// Mitsubishi GX Works2 project: 11国轩烘烤线体修改1028   PLC: Q06UDEH (continued)

lifter11203(ShuttleCarInOut:=LifterIO11203);(*出口升降台*)
LifterIO11203.xCylinder:=1;
Y246:=LifterIO11203.xCW;
Y247:=LifterIO11203.xCCW;
LifterIO11203.xForward:=M550;
LifterIO11203.xBackward:=M551;
ShuttleCarCurrentPosition(X51 OR X50,X50,X51,FALSE,LifterIO11203.iCurrentPos);
F455:=LifterIO11203.xOvertimeAlarm ;
LifterIO11203.diDeviceID:=11203;

Cylinder112011(ShuttleCarInOut:=	CylinderIO112011);	(*升降门*)
CylinderIO112011.xCylinder:=1;
Y240:=CylinderIO112011.xCW;(*修改*)				
Y241:=CylinderIO112011.xCCW;(*修改*)					
CylinderIO112011.xForward:=M556;				
CylinderIO112011.xBackward:=M557;				
ShuttleCarCurrentPosition(X4B OR X4A,X4B,X4A,FALSE,CylinderIO112011.iCurrentPos);				
F460:=CylinderIO112011.xOvertimeAlarm ;				
CylinderIO112011.diDeviceID:=112011;

Cylinder112012(ShuttleCarInOut:=	CylinderIO112012);	(*升降门*)
CylinderIO112012.xCylinder:=1;
Y242:=CylinderIO112012.xCW;	(*修改*)				
Y243:=CylinderIO112012.xCCW;		(*修改*)			
CylinderIO112012.xForward:=M558;				
CylinderIO112012.xBackward:=M559;				
ShuttleCarCurrentPosition(X4D OR X4C,X4D,X4C,FALSE,CylinderIO112012.iCurrentPos);				
F461:=CylinderIO112012.xOvertimeAlarm ;				
CylinderIO112012.diDeviceID:=112012;

Cylinder112041(ShuttleCarInOut:=	CylinderIO112041);	(*升降门*)
CylinderIO112041.xCylinder:=1;
Y24A:=CylinderIO112041.xCW;				
Y24B:=CylinderIO112041.xCCW;				
CylinderIO112041.xForward:=M560;				
CylinderIO112041.xBackward:=M561;				
ShuttleCarCurrentPosition(X54 OR X55,X55,X54,FALSE,CylinderIO112041.iCurrentPos);				
F462:=CylinderIO112041.xOvertimeAlarm ;				
CylinderIO112041.diDeviceID:=112041;

Cylinder112042(ShuttleCarInOut:=	CylinderIO112042);	(*升降门*)
CylinderIO112042.xCylinder:=1;
Y248:=CylinderIO112042.xCW;				
Y249:=CylinderIO112042.xCCW;				
CylinderIO112042.xForward:=M562;				
CylinderIO112042.xBackward:=M563;				
ShuttleCarCurrentPosition(X53 OR X52,X53,X52,FALSE,CylinderIO112042.iCurrentPos);				
F463:=CylinderIO112042.xOvertimeAlarm ;				
CylinderIO112042.diDeviceID:=112042;
	
Switch11301(ConveyorEntryIO:=	ConveyorIO111041,ConveyorExitIO:=	ConveyorIO11103,SwitchIO:=	SwitchIO11301);(*这里的Exit是为出线体，Entry为进线体*)
SwitchIO11301.xLiftCylinderRetractDetect:=X61;				
SwitchIO11301.xLiftCylinderExtendDetect:=X60;				
Y24C:=SwitchIO11301.xLiftCylinderExtend;				
SwitchIO11301.xLiftCylinderExtendButton:=M564;
SwitchIO11301.xLiftCylinderRetractButton:= NOT M564;		
F464:=SwitchIO11301.xOvertimeAlarm ;				

Switch11302(ConveyorEntryIO:= 	ConveyorIO111042,ConveyorExitIO:= 	ConveyorIO11106,SwitchIO:=	SwitchIO11302);
SwitchIO11302.xLiftCylinderRetractDetect:=X63;				
SwitchIO11302.xLiftCylinderExtendDetect:=X62;				
Y24D:=SwitchIO11302.xLiftCylinderExtend;				
SwitchIO11302.xLiftCylinderExtendButton:=M567;
SwitchIO11302.xLiftCylinderRetractButton:=NOT M567;				
F465:=SwitchIO11302.xOvertimeAlarm ;				

IF  m_i11315Task=1
  THEN 
 			Switch11315(ConveyorEntryIO:=ConveyorIO11137,ConveyorExitIO:=               ConveyorIO111381,	SwitchIO:= 	SwitchIO11315 );
   ELSE
     		Switch11315(ConveyorEntryIO:=ConveyorIO111381,ConveyorExitIO:=               ConveyorIO11137,	SwitchIO:= 	SwitchIO11315 );
END_IF;
SwitchIO11315.xLiftCylinderRetractDetect:=X7D;				
SwitchIO11315.xLiftCylinderExtendDetect:=X7C;				
Y25A:=SwitchIO11315.xLiftCylinderExtend;				
Y266:=SwitchIO11315.xEntryBarCylinderRetract;				
Y260:=(g_xAuto AND  m_i11315Task=2 )OR (M720 AND g_xManual) ;	(*十字路口阻挡气缸输出1*)	
Y261:=(g_xAuto AND  m_i11315Task=1 )OR ( M721 AND g_xManual);	(*十字路口阻挡气缸输出2*)
SwitchIO11315.xLiftCylinderExtendButton:=M568;	
SwitchIO11315.xLiftCylinderRetractButton:= NOT M568;	
SwitchIO11315.xEntryBarCylinderRetractButton:=M569;				
SwitchIO11315.xExitBarCylinderRetractButton:=M570;				
F466:=SwitchIO11315.xOvertimeAlarm ;				

Switch11316(ConveyorEntryIO:=ConveyorIO11140,ConveyorExitIO:= 	ConveyorIO111382,SwitchIO:= 	SwitchIO11316 );
SwitchIO11316.xLiftCylinderRetractDetect:=X7F;				
SwitchIO11316.xLiftCylinderExtendDetect:=X7E;				
Y25B:=SwitchIO11316.xLiftCylinderExtend;				
Y268:=NOT (m_i11316Task=2 OR M722);(*316阻挡气缸1*)		
Y269:=NOT (m_i11316Task=1 OR M723);	(*316阻挡气缸2*)	
SwitchIO11316.xLiftCylinderExtendButton:=M571;
SwitchIO11316.xLiftCylinderRetractButton:= NOT M571;				
SwitchIO11316.xEntryBarCylinderRetractButton:=M572;				
F467:=SwitchIO11316.xOvertimeAlarm ;				

UConveyor11303(	ConveyorIOLeft:=ConveyorIO11118,	ConveyorIORight:=ConveyorIO11120,	
									ConveyorIODown:=ConveyorIO11113,	UConveyorIO:=UConveyorIO11303);
UConveyorIO11303.xLiftCylinderExtendDetect1:=X64;
UConveyorIO11303.xLiftCylinderRetractDetect1:=X65;									
Y24E:=UConveyorIO11303.xLiftCylinderExtend1;								
Y262:=UConveyorIO11303.xExitBarCylinderRetract1;								
UConveyorIO11303.xLiftCylinderRetractDetect2:=X69;								
UConveyorIO11303.xLiftCylinderExtendDetect2:=X68;		
UConveyorIO11303.xBatteryDetect1:=X1A;		
Y250:=UConveyorIO11303.xLiftCylinderExtend2;								
UConveyorIO11303.xLiftCylinderExtendButton1:=M573;								
UConveyorIO11303.xExitBarCylinderRetractButton1:=M574;								
UConveyorIO11303.xLiftCylinderExtendButton2:=M575;								
F468:=UConveyorIO11303.xOvertimeAlarm ;								
(**X1A为电池检测保护*)

UConveyor11306(	ConveyorIOLeft:=ConveyorIO11121,	ConveyorIORight:=ConveyorIO11123,	
									ConveyorIODown:=ConveyorIO11114,	UConveyorIO:=UConveyorIO11306);
UConveyorIO11306.xLiftCylinderExtendDetect1:=X6A;	
UConveyorIO11306.xLiftCylinderRetractDetect1:=X6B;		
UConveyorIO11306.xBatteryDetect1:=X1F;							
Y251:=UConveyorIO11306.xLiftCylinderExtend1;								
Y263:=  UConveyorIO11306.xExitBarCylinderRetract1 ;								
UConveyorIO11306.xLiftCylinderRetractDetect2:=X6F;								
UConveyorIO11306.xLiftCylinderExtendDetect2:=X6E;								
Y253:=UConveyorIO11306.xLiftCylinderExtend2;								
UConveyorIO11306.xLiftCylinderExtendButton1:=M576;								
UConveyorIO11306.xExitBarCylinderRetractButton1:=M577;								
UConveyorIO11306.xLiftCylinderExtendButton2:=M578;								
F469:=UConveyorIO11306.xOvertimeAlarm ;								
(**X1F为电池检测保护*)

UConveyor11309(	ConveyorIOLeft:=ConveyorIO11124,	ConveyorIORight:=ConveyorIO11126,	
									ConveyorIODown:=ConveyorIO11115,	UConveyorIO:=UConveyorIO11309);
UConveyorIO11309.xLiftCylinderExtendDetect1:=X70;	
UConveyorIO11309.xLiftCylinderRetractDetect1:=X71;							
Y254:=UConveyorIO11309.xLiftCylinderExtend1;								
Y264:=UConveyorIO11309.xExitBarCylinderRetract1;								
UConveyorIO11309.xLiftCylinderRetractDetect2:=X75;								
UConveyorIO11309.xLiftCylinderExtendDetect2:=X74;								
Y256:=UConveyorIO11309.xLiftCylinderExtend2;								
UConveyorIO11309.xLiftCylinderExtendButton1:=M579;								
UConveyorIO11309.xExitBarCylinderRetractButton1:=M580;								
UConveyorIO11309.xLiftCylinderExtendButton2:=M581;								
F470:=UConveyorIO11309.xOvertimeAlarm ;								
(**X22为电池检测保护*)

UConveyor11312(	ConveyorIOLeft:=ConveyorIO11127,	ConveyorIORight:=ConveyorIO11129,	
									ConveyorIODown:=ConveyorIO11116,	UConveyorIO:=UConveyorIO11312);
UConveyorIO11312.xLiftCylinderExtendDetect1:=X76;
UConveyorIO11312.xLiftCylinderRetractDetect1:=X77;								
Y257:=UConveyorIO11312.xLiftCylinderExtend1;								
Y265:=UConveyorIO11312.xExitBarCylinderRetract1;								
UConveyorIO11312.xLiftCylinderRetractDetect2:=X7B;								
UConveyorIO11312.xLiftCylinderExtendDetect2:=X7A;								
Y259:=UConveyorIO11312.xLiftCylinderExtend2;								
UConveyorIO11312.xLiftCylinderExtendButton1:=M582;								
UConveyorIO11312.xExitBarCylinderRetractButton1:=M583;								
UConveyorIO11312.xLiftCylinderExtendButton2:=M584;								
F471:=UConveyorIO11312.xOvertimeAlarm ;								

(**************通信地址分配***************)
ComConveyor11104(ConveyorIO:=ConveyorIO11104,CommunicationIO:=ComConveyorIO11104);
ComCOnveyorIO11104.i_iResponsPCPLC:=D2001;	
ComCOnveyorIO11104.i_iReadWriteFlagPCPLC:=D2006;	
ComCOnveyorIO11104.i_iTaskProcessFlagPCPLC:=D2007;	
ComCOnveyorIO11104.i_iCommandPCPLC:=D2008;	
ComCOnveyorIO11104.i_iTaskIDPCPLC:=D2009;	
DMOV(TRUE,D2010,ComConveyorIO11104.i_diDestinationDevicePCPLC);	
ComCOnveyorIO11104.i_iProductIDPCPLC:=D2012;	
D3001:=ComCOnveyorIO11104.o_iRequestPLCPC;	
D3006:=ComCOnveyorIO11104.o_iReadWriteFlagPLCPC;	
D3007:=ComCOnveyorIO11104.o_iDeviceStatusPLCPC;	
D3008:=ComCOnveyorIO11104.o_iTaskIDPLCPC;	
D3009:=ComCOnveyorIO11104.o_iProductIDPLCPC;	

ComConveyor11108(ConveyorIO:=ConveyorIO11108,CommunicationIO:=ComConveyorIO11108);
ComCOnveyorIO11108.i_iResponsPCPLC:=D2016;	
ComCOnveyorIO11108.i_iReadWriteFlagPCPLC:=D2021;	
ComCOnveyorIO11108.i_iTaskProcessFlagPCPLC:=D2022;	
ComCOnveyorIO11108.i_iCommandPCPLC:=D2023;	
ComCOnveyorIO11108.i_iTaskIDPCPLC:=D2024;	
DMOV(TRUE,D2025,ComConveyorIO11108.i_diDestinationDevicePCPLC);		
ComCOnveyorIO11108.i_iProductIDPCPLC:=D2027;	
D3016:=ComCOnveyorIO11108.o_iRequestPLCPC;	
D3021:=ComCOnveyorIO11108.o_iReadWriteFlagPLCPC;	
D3022:=ComCOnveyorIO11108.o_iDeviceStatusPLCPC;	
D3023:=ComCOnveyorIO11108.o_iTaskIDPLCPC;	
D3024:=ComCOnveyorIO11108.o_iProductIDPLCPC;	

ComConveyor11107(ConveyorIO:=ConveyorIO11107,CommunicationIO:=ComConveyorIO11107);
ComConveyorIO11107.i_iResponsPCPLC:=D2031;	
ComConveyorIO11107.i_iReadWriteFlagPCPLC:=D2036;	
ComConveyorIO11107.i_iTaskProcessFlagPCPLC:=D2037;	
ComConveyorIO11107.i_iCommandPCPLC:=D2038;	
ComConveyorIO11107.i_iTaskIDPCPLC:=D2039;	
DMOV(TRUE,D2040,ComConveyorIO11107.i_diDestinationDevicePCPLC);	
ComConveyorIO11107.i_iProductIDPCPLC:=D2042;	
D3031:=ComConveyorIO11107.o_iRequestPLCPC;	
D3036:=ComConveyorIO11107.o_iReadWriteFlagPLCPC;	
D3037:=ComConveyorIO11107.o_iDeviceStatusPLCPC;	
D3038:=ComConveyorIO11107.o_iTaskIDPLCPC;	
D3039:=ComConveyorIO11107.o_iProductIDPLCPC;	
	

ComConveyor11142(ConveyorIO:=ConveyorIO11142,CommunicationIO:=ComConveyorIO11142);
ComCOnveyorIO11142.i_iResponsPCPLC:=D2046;	
ComCOnveyorIO11142.i_iReadWriteFlagPCPLC:=D2051;	
ComCOnveyorIO11142.i_iTaskProcessFlagPCPLC:=D2052;	
ComCOnveyorIO11142.i_iCommandPCPLC:=D2053;	
ComCOnveyorIO11142.i_iTaskIDPCPLC:=D2054;	
DMOV(TRUE,D2055,ComConveyorIO11142.i_diDestinationDevicePCPLC);	
ComCOnveyorIO11142.i_iProductIDPCPLC:=D2057;	
D3046:=ComCOnveyorIO11142.o_iRequestPLCPC;	
D3051:=ComCOnveyorIO11142.o_iReadWriteFlagPLCPC;	
D3052:=ComCOnveyorIO11142.o_iDeviceStatusPLCPC;	
D3053:=ComCOnveyorIO11142.o_iTaskIDPLCPC;	
D3054:=ComCOnveyorIO11142.o_iProductIDPLCPC;	

ComConveyor11141(ConveyorIO:=ConveyorIO11141,CommunicationIO:=ComConveyorIO11141);
ComCOnveyorIO11141.i_iResponsPCPLC:=D2061;	
ComCOnveyorIO11141.i_iReadWriteFlagPCPLC:=D2066;	
ComCOnveyorIO11141.i_iTaskProcessFlagPCPLC:=D2067;	
ComCOnveyorIO11141.i_iCommandPCPLC:=D2068;	
ComCOnveyorIO11141.i_iTaskIDPCPLC:=D2069;	
DMOV(TRUE,D2070,ComConveyorIO11141.i_diDestinationDevicePCPLC);	
ComCOnveyorIO11141.i_iProductIDPCPLC:=D2072;	
D3061:=ComCOnveyorIO11141.o_iRequestPLCPC;	
D3066:=ComCOnveyorIO11141.o_iReadWriteFlagPLCPC;	
D3067:=ComCOnveyorIO11141.o_iDeviceStatusPLCPC;	
D3068:=ComCOnveyorIO11141.o_iTaskIDPLCPC;	
D3069:=ComCOnveyorIO11141.o_iProductIDPLCPC;	

ComConveyor11110(ConveyorIO:=ConveyorIO11110,CommunicationIO:=ComConveyorIO11110);
ComCOnveyorIO11110.i_iResponsPCPLC:=D2076;	
ComCOnveyorIO11110.i_iReadWriteFlagPCPLC:=D2081;	
ComCOnveyorIO11110.i_iTaskProcessFlagPCPLC:=D2082;	
ComCOnveyorIO11110.i_iCommandPCPLC:=D2083;	
ComCOnveyorIO11110.i_iTaskIDPCPLC:=D2084;	
DMOV(TRUE,D2085,ComConveyorIO11110.i_diDestinationDevicePCPLC);	
ComCOnveyorIO11110.i_iProductIDPCPLC:=D2087;	
D3076:=ComCOnveyorIO11110.o_iRequestPLCPC;	
D3081:=ComCOnveyorIO11110.o_iReadWriteFlagPLCPC;	
D3082:=ComCOnveyorIO11110.o_iDeviceStatusPLCPC;	
D3083:=ComCOnveyorIO11110.o_iTaskIDPLCPC;	
D3084:=ComCOnveyorIO11110.o_iProductIDPLCPC;	

ComConveyor11111(ConveyorIO:=ConveyorIO11111,CommunicationIO:=ComConveyorIO11111);
ComCOnveyorIO11111.i_iResponsPCPLC:=D2091;	
ComCOnveyorIO11111.i_iReadWriteFlagPCPLC:=D2096;	
ComCOnveyorIO11111.i_iTaskProcessFlagPCPLC:=D2097;	
ComCOnveyorIO11111.i_iCommandPCPLC:=D2098;	
ComCOnveyorIO11111.i_iTaskIDPCPLC:=D2099;	
DMOV(TRUE,D2100,ComConveyorIO11111.i_diDestinationDevicePCPLC);	
ComCOnveyorIO11111.i_iProductIDPCPLC:=D2102;	
D3091:=ComCOnveyorIO11111.o_iRequestPLCPC;	
D3096:=ComCOnveyorIO11111.o_iReadWriteFlagPLCPC;	
D3097:=ComCOnveyorIO11111.o_iDeviceStatusPLCPC;	
D3098:=ComCOnveyorIO11111.o_iTaskIDPLCPC;	
D3099:=ComCOnveyorIO11111.o_iProductIDPLCPC;	

ComConveyor11143(ConveyorIO:=ConveyorIO11143,CommunicationIO:=ComConveyorIO11143);
ComConveyorIO11143.i_iResponsPCPLC:=D2106;	
ComConveyorIO11143.i_iReadWriteFlagPCPLC:=D2111;	
ComConveyorIO11143.i_iTaskProcessFlagPCPLC:=D2112;	
ComConveyorIO11143.i_iCommandPCPLC:=D2113;	
ComConveyorIO11143.i_iTaskIDPCPLC:=D2114;	
DMOV(TRUE,D2115,ComConveyorIO11143.i_diDestinationDevicePCPLC);	
ComConveyorIO11143.i_iProductIDPCPLC:=D2117;	
D3106:=ComConveyorIO11143.o_iRequestPLCPC;	
D3111:=ComConveyorIO11143.o_iReadWriteFlagPLCPC;	
D3112:=ComConveyorIO11143.o_iDeviceStatusPLCPC;	
D3113:=ComConveyorIO11143.o_iTaskIDPLCPC;	
D3114:=ComConveyorIO11143.o_iProductIDPLCPC;	

(*///////////////////////////////////自动部分/////////////////////////////*)
IF g_xAuto    THEN
			(*门直接用Y控制，不用块了*)
			CylinderIO112011.xMDIExe:=1;
		IF D401.2  AND 	ConveyorIO11101.xEmpty  AND CylinderIO112012.iCurrentPos=1
			THEN(*上层10给11有料信号401.2*)
						CylinderIO112011.iDestinationPos:=2;
			ELSE CylinderIO112011.iDestinationPos:=1; (*如果10有下料信号但是11对接线体也有料，则关闭AB门*)
		END_IF;	
		D201.2:=CylinderIO112011.iCurrentPos=2 AND ConveyorIO11101.xEmpty;(*11给10的上层下料允许对接信号*)
		ConveyorIO11101.xLoad:=D401.4;(*10线体的下料信号*)
		(*第2个隔离门*)
		CylinderIO112012.xMDIExe:=1;
		IF NOT ConveyorIO11101.xEmpty  AND CylinderIO112011.iCurrentPos=1 (*第二个隔离门只有在第一个隔离门关住后*)
			THEN
							CylinderIO112012.iDestinationPos:=2;
			ELSE 	CylinderIO112012.iDestinationPos:=1;
		END_IF;		
		ConveyorIO11101.xUnload:=ConveyorIO11102.xEmpty AND CylinderIO112012.iCurrentPos=2;
		ConveyorIO11102.xLoad:=ConveyorIO11101.xNextRun;
		Switch11301Task(xCondition:= Switch11301Condition,(*抢占排队*)
									xTaskComplete:=LDP(TRUE,ConveyorIO111041.xEmpty) ,
									xReset:=g_diDeviceIDSelect=11104 AND g_xResetSingle ,
									iPriority:=m_i11301Task);
		Switch11301Condition[1]:=ConveyorIO11102.xEmpty=0 AND ConveyorIO11104.xEmpty;(*顶升移栽任务1,往烘烤*)
		Switch11301Condition[2]:=ConveyorIO11109.xEmpty=0 AND ConveyorIO11111.xEmpty AND LifterIO11202.iCurrentPos=2;(*顶升移栽任务2，往机械手*)
		ConveyorIO11102.xUnload:=ConveyorIO111041.xEmpty AND m_i11301Task=1;
		SwitchIO11301.xLiftCylinderExtendInit:=1;(*初始化顶起*)
		SwitchIO11301.xEntryEnable:=ConveyorIO11102.xNextRun;
		SwitchIO11301.xSwithEnable:=m_i11301Task=2;(*任务2要直行，降下气缸*)
		SwitchIO11301.xExitEnable:=(ConveyorIO11104.xEmpty AND m_i11301Task=1)(*1041虚拟线体运给104*)
													OR(ConveyorIO11111.xEmpty AND m_i11301Task=2);(*11103出料给11111*)
		(*满框去烘烤*)													
		ConveyorIO11104.xLoad:=ConveyorIO111041.xNextRun;
		ConveyorIO11104.xUnload:=ConveyorIO111042.xEmpty;(*这里到时候需要加一个扫码条件，判断去哪个烘烤库*)
		SwitchIO11302.xEntryEnable:=ConveyorIO11104.xNextRun;
		SwitchIO11302.xSwithEnable:=1;
		SwitchIO11302.xLiftCylinderExtendInit:=1;(*初始化顶起*)
		SwitchIO11302.xExitEnable:=(ConveyorIO111042.diDesConveyor=11108 AND ConveyorIO11108.xEmpty)
													OR (ConveyorIO111042.diDesConveyor=11107 AND ConveyorIO11107.xEmpty);
		ConveyorIO11106.xUnloadCCW:=ConveyorIO111042.diDesConveyor=11108;
		ConveyorIO11107.xLoad:=ConveyorIO11106.xNextRun AND  ConveyorIO11106.diDesConveyor=11107;
		ConveyorIO11108.xLoad:=ConveyorIO11106.xNextRun AND ConveyorIO11106.diDesConveyor=11108;
		(*未增加11107和11108下料信号，与工控机信号对接*)
		Switch11316Task(arrxCondition:=Switch11316Condition ,
								xTaskComplete:= LDF(TRUE,ConveyorIO11138.xEmpty),
								xReset:= g_xResetSingle AND g_diDeviceIDSelect=11138,	
								iPriority:=m_i11316Task);
		Switch11316Condition[1].xCondition:=ConveyorIO11141.xEmpty=0;
		Switch11316Condition[2].xCondition:=ConveyorIO11142.xEmpty=0;
		
		LifterIO11204.xMDIExe:=NOT ConveyorIO11140.xError AND NOT ConveyorIO11141.xError ;
		IF NOT ConveyorIO11142.xEmpty   THEN
			LifterIO11204.iDestinationPos:=1;
		ELSE 
			LifterIO11204.iDestinationPos:=2;
		END_IF;	

		LifterIO11205.xMDIExe:=NOT ConveyorIO11140.xError AND NOT ConveyorIO11142.xError ;
		IF NOT ConveyorIO11141.xEmpty THEN
			LifterIO11205.iDestinationPos:=1;
		ELSE
			LifterIO11205.iDestinationPos:=2;
		END_IF;	
		
		(*ConveyorIO11141.xPutInto:=  M880;*)(*这里需要上位机给命令，以后需要就加*)
	(*	ConveyorIO11142.xPutInto:=  M881;*)(*这里需要上位机给命令，以后需要就加*)
		ConveyorIO11141.xUnload:=ConveyorIO11140.xEmpty AND m_i11316Task=1 ; (*AND LifterIO11204.iCurrentPos=1;*)(*这里可能需要Load，接到堆垛机指令就Load，以后需要就加*)
		ConveyorIO11142.xUnload:=ConveyorIO11140.xEmpty AND m_i11316Task=2;(*  AND LifterIO11205.iCurrentPos=1;*)
		SwitchIO11316.xEntryEnable:=(ConveyorIO11141.xNextRun AND m_i11316Task=1)
													OR (ConveyorIO11142.xNextRun AND m_i11316Task=2);
		ConveyorIO11140.xloadCCW:= m_i11316Task=1;													
		SwitchIO11316.xSwithEnable:=1;
		SwitchIO11316.xExitEnable:=ConveyorIO11138.xEmpty;
		(*下层十字路口——+——+——+——+——+——+——+——+——+——+*)
		Switch11315Task(xCondition:=Switch11315Condition ,
									xTaskComplete:=LDF(TRUE,(ConveyorIO11109.xEmpty AND m_i11315Task=2 )OR(ConveyorIO11143.xEmpty AND m_i11315Task=1) ),
									xReset:=g_xResetSingle AND g_diDeviceIDSelect=11138 ,
									iPriority:= m_i11315Task );
		Switch11315Condition[1]:=ConveyorIO11136.xEmpty=0 AND ConveyorIO11143.xEmpty;
		Switch11315Condition[2]:=(ConveyorIO11140.xEmpty=0 OR ConveyorIO111382.xEmpty=0) AND ConveyorIO11109.xEmpty AND LifterIO11202.iCurrentPos=1;(*像这种带位置判断的，最好把检测开关也加上去*)
		SwitchIO11315.xEntryEnable:=ConveyorIO11136.xNextRun OR ConveyorIO11138.xNextRun ;
		SwitchIO11315.xSwithEnable:=(*m_i11315Task=1 *)1 ;
		SwitchIO11315.xExitEnable:=(m_i11315Task=1 AND  ConveyorIO11143.xEmpty)
													OR (m_i11315Task=2 AND ConveyorIO11109.xEmpty AND  LifterIO11202.iCurrentPos=1);
		ConveyorIO11138.xload:=ConveyorIO111382.xNextRun;
		ConveyorIO11138.xUnload:=ConveyorIO111381.xEmpty AND m_i11315Task=2 AND SwitchIO11315.xLiftCylinderExtendDetect  ;
		ConveyorIO11109.xLoad:=ConveyorIO11137.xNextRun AND m_i11315Task =2;

		IF m_i11315Task=2 THEN(*任务2时，升降由11137的状态控制，1时会由Switch块自己控制。因为任务2时，走134的step,不会控制升降*)
(*			IF NOT ConveyorIO11138.xEmpty THEN
				SwitchIO11315.xLiftCylinderExtend:=1;
				SwitchIO11315.xLiftCylinderRetract:=0;
			ELSE
				SwitchIO11315.xLiftCylinderExtend:=0;
				SwitchIO11315.xLiftCylinderRetract:=1;	
			END_IF;*)
			SwitchIO11315.xLiftCylinderExtendInit:=1;
		ELSE
			SwitchIO11315.xLiftCylinderExtendInit:=0;
		END_IF;
	

		IF LDP(TRUE,NOT ConveyorIO111381.xEmpty )THEN(*原来136和137公用一个光电检测开关，137竖向，136横向，当137有料时136也有料，这里用来给136直接下料，修改后用于1381虚拟线体和137线体*)
	ConveyorIO11137.xPutInto:=1;
		ELSIF	 LDP(TRUE,NOT ConveyorIO11137.xEmpty )THEN
			ConveyorIO11137.xPutInto:=0;
		END_IF;	

													
(*11202升降控制*)
													
		LifterIO11202.xMDIExe:=NOT ConveyorIO11109.xError AND NOT ConveyorIO11103.xError AND NOT ConveyorIO11137.xError;
		ConveyorIO11109.xloadCCW:=1;
		IF ConveyorIO11109.xEmpty THEN
			LifterIO11202.iDestinationPos:=1;
		ELSE
			LifterIO11202.iDestinationPos:=2;
		END_IF;	
		IF m_i11301Task=2 THEN
		SwitchIO11301.xLiftCylinderExtend:=0;
		SwitchIO11301.xLiftCylinderRetract:=1;
		END_IF;	 
		ConveyorIO11109.xUnload:=ConveyorIO11103.xEmpty AND LifterIO11202.iCurrentPos=2 AND m_i11301Task=2;
		ConveyorIO11103.xLoad:=ConveyorIO11109.xNextRun;
		IF LDP(TRUE,ConveyorIO11103.xEmpty=0) AND m_i11301Task=2 THEN
			ConveyorIO111041.xPutInto:=1;
		ELSIF LDP(TRUE,ConveyorIO111041.xEmpty=0) AND m_i11301Task=2 THEN
			ConveyorIO111041.xPutInto:=0;	
		END_IF;
		(*烘烤出去机械手*)
		ConveyorIO11111.xLoad:=ConveyorIO11103.xNextRun;
		ConveyorIO11111.xUnload:=ConveyorIO11112.xEmpty;
		ConveyorIO11112.xLoad:=ConveyorIO11111.xNextRun;
		ConveyorIO11112.xUnload:=ConveyorIO11105.xEmpty;
		ConveyorIO11105.xLoad:=ConveyorIO11112.xNextRun;
		ConveyorIO11105.xUnload:=ConveyorIO11139.xEmpty;
		ConveyorIO11139.xLoad:=ConveyorIO11105.xNextRun;
		ConveyorIO11139.xUnload:=UConveyorio11303.iTask=1 AND m_xU1TaskStart;(*39下料给U1*)


		Conveyor11139Task(arrxCondition:=Conveyor11139Condition,
											xTaskComplete:=LDP(TRUE,ConveyorIO11139.xEmpty),
											xReset:= g_xResetSingle AND g_diDeviceIDSelect=11139 ,
											iPriority:= m_i11139Task);
		Conveyor11139Condition[1].xCondition:=ConveyorIO111181.xEmpty AND m_xLoadPermit1;
		Conveyor11139Condition[2].xCondition:=ConveyorIO111231.xEmpty  AND m_xLoadPermit2;
		Conveyor11139Condition[3].xCondition:=ConveyorIO111241.xEmpty  AND m_xLoadPermit3;
		Conveyor11139Condition[4].xCondition:=ConveyorIO111291.xEmpty  AND m_xLoadPermit4; 
		DMOV(m_i11139Task=1,	11118,	ConveyorIO11139.diDesConveyor);(*上电时，机械手U型线体处空时生成任务号，并进行抢占*)
		DMOV(m_i11139Task=2,	11123,	ConveyorIO11139.diDesConveyor);
		DMOV(m_i11139Task=3,	11124,	ConveyorIO11139.diDesConveyor);
		DMOV(m_i11139Task=4,	11129,	ConveyorIO11139.diDesConveyor);

		(*这个PickDone信号，他们给信号时置位，为empty的上升沿复位*)
		SET(XA0	AND NOT ConveyorIO11119.xEmpty,	m_xPickDone[1]);	
		RST(ConveyorIO11119.xEmpty,	m_xPickDone[1]);
		SET(XA1 	AND NOT ConveyorIO11122.xEmpty,	m_xPickDone[2]);	
		RST(ConveyorIO11122.xEmpty,	m_xPickDone[2]);
		SET(XA2	AND NOT ConveyorIO11125.xEmpty,	m_xPickDone[3]);	
		RST(ConveyorIO11125.xEmpty,	m_xPickDone[3]);
		SET(XA3	AND NOT ConveyorIO11128.xEmpty,	m_xPickDone[4]);	
		RST(ConveyorIO11128.xEmpty,	m_xPickDone[4]);

		DMOV(m_xPickDone[1] AND ConveyorIO11145.xEmpty AND ConveyorIO11145.diDesConveyor=0,	11117,	ConveyorIO11145.diDesConveyor);(*机械手给空框完成信号后将提升机线体作为目标地址发送，空框一直送至11117*)
		DMOV(m_xPickDone[2] AND ConveyorIO11146.xEmpty AND ConveyorIO11146.diDesConveyor=0,	11117,	ConveyorIO11146.diDesConveyor);
		DMOV(m_xPickDone[3] AND ConveyorIO11147.xEmpty AND ConveyorIO11147.diDesConveyor=0,	11117,	ConveyorIO11147.diDesConveyor);
		DMOV(m_xPickDone[4],	11117,	ConveyorIO11128.diDesConveyor);(*最初始的目标地址生成,*)

		(*目标地址的传递，横纵传递分开写，横纵之间的传递在块里写好了，不用担心*)
		ConveyorIO11113.diDesConveyorIn:=	ConveyorIO11139.diDesConveyorOut;
		ConveyorIO11145.diDesConveyorIn:=	ConveyorIO11113.diDesConveyorOut;
		ConveyorIO11114.diDesConveyorIn:=	ConveyorIO11145.diDesConveyorOut;
		ConveyorIO11146.diDesConveyorIn:=	ConveyorIO11114.diDesConveyorOut;
		ConveyorIO11115.diDesConveyorIn:=	ConveyorIO11146.diDesConveyorOut;
		ConveyorIO11147.diDesConveyorIn:=	ConveyorIO11115.diDesConveyorOut;
		ConveyorIO11116.diDesConveyorIn:=	ConveyorIO11147.diDesConveyorOut;
		(*纵向任务传递，包括虚拟线体*)
		ConveyorIO11120.diDesConveyorIn:=	ConveyorIO11119.diDesConveyorOut;
		ConveyorIO11121.diDesConveyorIn:=	ConveyorIO11122.diDesConveyorOut;
		ConveyorIO11126.diDesConveyorIn:=	ConveyorIO11125.diDesConveyorOut;
		ConveyorIO11127.diDesConveyorIn:=	ConveyorIO11128.diDesConveyorOut;
		ConveyorIO111042.diDesConveyor:=11107;


		m_TPU1TaskComplete(IN:=ConveyorIO11113.xEmpty ,PT:=t#200ms,Q:= m_xU1TaskComplete,ET:= m_tU1TaskComplete );
		m_TonU1TaskStart(IN:= ConveyorIO11113.xEmpty ,PT:= t#300MS ,Q:=m_xU1TaskStart ,ET:=m_tU1TaskStart );
		Uconveyor11303Task(xCondition:=Uconveyor11303Condition,
											xTaskComplete:=LDF(TRUE,m_xU1TaskComplete) ,
											xReset:= g_xResetSingle AND g_diDeviceIDSelect=11113 ,
											iPriority:=UConveyorio11303.iTask );
			Uconveyor11303Condition[1]:=ConveyorIO11139.xEmpty=0 AND m_i11139Task>0;(*这里还要再改的*)(*任务1是U块入料到机械手*)
			Uconveyor11303Condition[3]:=ConveyorIO111201.xEmpty=0  AND m_xPickDone[1];	(*任务3是右臂出料*)
		UConveyorio11303.xEntryEnable1:=ConveyorIO11139.xNextRun;(*U型横向线体入料使能，EntryEnable1，2，3都是在任务1时用*)
		UConveyorIO11303.xEntryEnable3:=ConveyorIO111201.xNextRun;(*U型右臂入料使能*)
		UConveyorio11303.xExitEnable1:=ConveyorIO11145.xEmpty ;(*xExitEnable1是主线体出，2是左臂出，3是右臂出，这个为横向线体出料使能*)
		UConveyorio11303.xExitEnable3:=ConveyorIO111181.xEmpty;(*这个为右臂出料使能*)
	
		ConveyorIO111181.xLoad:=ConveyorIO11118.xNextRun;(*这里是U块左右臂再增加一段线体时使用，用于控制该线体*)
		IF ConveyorIO111181.xEmpty=0  AND ConveyorIO11119.xEmpty THEN
			UConveyorIO11303.xLiftCylinderExtend2:=0;
			UConveyorIO11303.xLiftCylinderRetract2:=1;(*Extend2和Retract2为右臂顶升移栽气缸伸出和收回，Extend1和Retract1为左臂顶升移栽气缸伸出和收回*)
		END_IF;	
		ConveyorIO111181.xUnload:=ConveyorIO11119.xEmpty AND UConveyorIO11303.xLiftCylinderRetractDetect1 AND UConveyorIO11303.xLiftCylinderRetractDetect2;(*机械手横向线体控制*)
		ConveyorIO11119.xLoad:=ConveyorIO111181.xNextRun AND UConveyorIO11303.xLiftCylinderRetractDetect1 AND UConveyorIO11303.xLiftCylinderRetractDetect1;
			m_Ton11119(IN:= NOT ConveyorIO11119.xEmpty,PT:= t#3s ,Q:= m_x111201 ,ET:= m_t111201);
		IF NOT ConveyorIO11119.xEmpty AND m_x111201 THEN(*需加延时刷新111201，线体第0步要延时100ms才能检测有料，*)
			ConveyorIO111201.xPutInto:=1;
		ELSE 
			ConveyorIO111201.xPutInto:=0;
		END_IF;	
		ConveyorIO111201.xUnload:=ConveyorIO11120.xEmpty AND UConveyorio11303.iTask=3 ;(*右臂出料*)
	(**)	
		ConveyorIO11120.xLoadCCW:=1;
(*	 UConveyorIO11303.	xLiftCylinderExtendInit1=1 *)
		(*至此，U1的动作全部完成*)
		(*过度线体145*)
		ConveyorIO11145.xLoad:=ConveyorIO11113.xNextRun;
		ConveyorIO11145.xUnload:=(UConveyorio11306.iTask=1  AND m_xU2TaskStart )OR (ConveyorIO11146.diDesConveyor=11117 AND ConveyorIO11115.xEmpty) ;
		(*U2块*)
		m_TPU2TaskComplete(IN:=ConveyorIO11114.xEmpty ,PT:=t#200ms,Q:= m_xU2TaskComplete,ET:= m_tU2TaskComplete );
		m_TonU2TaskStart(IN:= ConveyorIO11114.xEmpty ,PT:= t#300MS ,Q:=m_xU2TaskStart ,ET:=m_tU2TaskStart );
		Uconveyor11306Task(xCondition:=Uconveyor11306Condition,
											xTaskComplete:=LDF(TRUE,m_xU2TaskComplete) ,
											xReset:= g_xResetSingle AND g_diDeviceIDSelect=11114,
											iPriority:=UConveyorIO11306.iTask );
			Uconveyor11306Condition[1]:=ConveyorIO11145.xEmpty=0 AND ConveyorIO11145.diDesConveyor<>11118
																														AND ConveyorIO11145.diDesConveyor<>0;(*这里还要再改的*)
			Uconveyor11306Condition[2]:=ConveyorIO111211.xEmpty=0  AND m_xPickDone[2];(*任务2是左臂出料*)
		UConveyorio11306.xEntryEnable1:=ConveyorIO11145.xNextRun ;
		UConveyorIO11306.xEntryEnable2:=ConveyorIO111211.xNextRun;
		UConveyorio11306.xExitEnable1:=ConveyorIO11146.xEmpty ;(*U型块任务1都是进前判断3个任务：往左进，往右进，主线体直接走，2是往左臂线体出，3是往右臂线体出*)
		UConveyorio11306.xExitEnable2:=ConveyorIO111231.xEmpty;(*xExitEnable1是主线体出，2是左臂出，3是右臂出*)
		ConveyorIO111231.xLoad:=ConveyorIO11123.xNextRun;

		IF ConveyorIO111231.xEmpty=0  AND ConveyorIO11122.xEmpty THEN
			UConveyorIO11306.xLiftCylinderExtend1:=0;
			UConveyorIO11306.xLiftCylinderRetract1:=1;(*U1,U3用2，U2,U4用1*)
		END_IF;	
		ConveyorIO111231.xUnload:=ConveyorIO11122.xEmpty AND UConveyorIO11306.xLiftCylinderRetractDetect1 AND UConveyorIO11306.xLiftCylinderRetractDetect2;(*机械手横向线体控制*)
		ConveyorIO11122.xLoad:=ConveyorIO111231.xNextRun AND UConveyorIO11306.xLiftCylinderRetractDetect1 AND UConveyorIO11306.xLiftCylinderRetractDetect2;
		m_Ton11122(IN:= NOT ConveyorIO11122.xEmpty,PT:= t#3s ,Q:= m_x111211 ,ET:= m_t111211);
		IF NOT ConveyorIO11122.xEmpty AND m_x111211 THEN(*加延时刷新111211，线体第0步要延时100ms才能检测有料，*)
			ConveyorIO111211.xPutInto:=1;
		ELSIF ConveyorIO111211.xEmpty=0 THEN
			ConveyorIO111211.xPutInto:=0;
		END_IF;	
		ConveyorIO111211.xUnload:=ConveyorIO11121.xEmpty AND UConveyorio11306.iTask=2 ;(*左臂下料*)
		(*至此，U2的动作全部完成*)
		(*过度线体146*)
		ConveyorIO11146.xLoad:=ConveyorIO11114.xNextRun;
		ConveyorIO11146.xUnload:=(UConveyorio11309.iTask=1 AND m_xU3TaskStart )OR (ConveyorIO11146.diDesConveyor=11117 AND ConveyorIO11115.xEmpty) ;
		(*U3块*)
		m_TPU3TaskComplete(IN:=ConveyorIO11115.xEmpty ,PT:=t#200ms,Q:= m_xU3TaskComplete,ET:= m_tU3TaskComplete );
		m_TonU3TaskStart(IN:= ConveyorIO11115.xEmpty ,PT:= t#300MS ,Q:=m_xU3TaskStart ,ET:=m_tU3TaskStart );
		Uconveyor11309Task(xCondition:=Uconveyor11309Condition,
											xTaskComplete:=LDF(TRUE,m_xU3TaskComplete) ,
											xReset:= g_xResetSingle AND g_diDeviceIDSelect=11115,
											iPriority:=UConveyorIO11309.iTask );
			Uconveyor11309Condition[1]:=ConveyorIO11146.xEmpty=0 AND ConveyorIO11146.diDesConveyor<>11123
																														AND ConveyorIO11146.diDesConveyor<>0;(*这里还要再改的*)
			Uconveyor11309Condition[3]:=ConveyorIO111261.xEmpty=0 AND m_xPickDone[3] ;	
		UConveyorio11309.xEntryEnable1:=ConveyorIO11146.xNextRun;
		UConveyorIO11309.xEntryEnable3:=ConveyorIO111261.xNextRun;

		UConveyorio11309.xExitEnable1:=ConveyorIO11147.xEmpty ;(*U型块任务1都是进前判断3个任务：往左进，往右进，主线体直接走，2是往左臂线体出，3是往右臂线体出*)
		UConveyorio11309.xExitEnable3:=ConveyorIO111241.xEmpty;(*xExitEnable1是主线体出，2是左臂出，3是右臂出*)
		ConveyorIO111241.xLoad:=ConveyorIO11124.xNextRun;

		IF ConveyorIO111241.xEmpty=0  AND ConveyorIO11125.xEmpty THEN
			UConveyorio11309.xLiftCylinderExtend2:=0;
			UConveyorio11309.xLiftCylinderRetract2:=1;(*U1,U3用2，U2,U4用1*)
		END_IF;	
		ConveyorIO111241.xUnload:=ConveyorIO11125.xEmpty AND UConveyorio11309.xLiftCylinderRetractDetect2 AND UConveyorio11309.xLiftCylinderRetractDetect1;(*机械手横向线体控制*)
		ConveyorIO11125.xLoad:=ConveyorIO111241.xNextRun AND UConveyorio11309.xLiftCylinderRetractDetect2 AND UConveyorio11309.xLiftCylinderRetractDetect1;
		m_Ton11125(IN:= NOT ConveyorIO11125.xEmpty,PT:= t#3s ,Q:= m_x111261 ,ET:= m_t111261);
		IF NOT ConveyorIO11125.xEmpty AND m_x111261 THEN(*加延时刷新111261，线体第0步要延时100ms才能检测有料，*)
			ConveyorIO111261.xPutInto:=1;
		ELSIF ConveyorIO111261.xEmpty=0 THEN
			ConveyorIO111261.xPutInto:=0;
		END_IF;	
				ConveyorIO111261.xUnload:=ConveyorIO11126.xEmpty AND UConveyorio11309.iTask=3 ;
		(*至此，U3的动作全部完成*)
		(*过度线体147*)
		ConveyorIO11147.xLoad:=ConveyorIO11115.xNextRun;
		ConveyorIO11147.xUnload:=(UConveyorio11312.iTask=1 AND m_xU4TaskStart) OR (ConveyorIO11147.diDesConveyor=11117 AND ConveyorIO11116.xEmpty) ;
		(*U4块*)
		m_TPU4TaskComplete(IN:=ConveyorIO11116.xEmpty ,PT:=t#200ms,Q:= m_xU4TaskComplete,ET:= m_tU4TaskComplete );
		m_TonU4TaskStart(IN:= ConveyorIO11116.xEmpty ,PT:= t#300MS ,Q:=m_xU4TaskStart ,ET:=m_tU4TaskStart );
		Uconveyor11312Task(xCondition:=Uconveyor11312Condition,
											xTaskComplete:=LDF(TRUE,m_xU4TaskComplete) ,
											xReset:= g_xResetSingle AND g_diDeviceIDSelect=11116,
											iPriority:=UConveyorIO11312.iTask );
			Uconveyor11312Condition[1]:=ConveyorIO11147.xEmpty=0 AND ConveyorIO11147.diDesConveyor<>11124
																														AND ConveyorIO11147.diDesConveyor<>0;(*这里还要再改的*)
	Uconveyor11312Condition[2]:=ConveyorIO11128.xEmpty=0  AND m_xPickDone[4] ;	
		UConveyorio11312.xEntryEnable1:=ConveyorIO11147.xNextRun;
		UConveyorIO11312.xEntryEnable2:=ConveyorIO111271.xNextRun;
		UConveyorio11312.xExitEnable1:=ConveyorIO11117.xEmpty AND  LifterIO11203.iCurrentPos=2;
		UConveyorio11312.xExitEnable2:=ConveyorIO111291.xEmpty;
		ConveyorIO111291.xLoad:=ConveyorIO11129.xNextRun;

		IF ConveyorIO111291.xEmpty=0  AND ConveyorIO11128.xEmpty THEN
			UConveyorio11312.xLiftCylinderExtend1:=0;
			UConveyorio11312.xLiftCylinderRetract1:=1;(*U1,U3用2，U2,U4用1*)
		END_IF;	
		ConveyorIO111291.xUnload:=ConveyorIO11128.xEmpty AND UConveyorio11312.xLiftCylinderRetractDetect1 AND UConveyorio11312.xLiftCylinderRetractDetect2;(*机械手横向线体控制*)
		ConveyorIO11128.xLoad:=ConveyorIO111291.xNextRun AND UConveyorio11312.xLiftCylinderRetractDetect1 AND UConveyorio11312.xLiftCylinderRetractDetect2;
		m_Ton11128(IN:= NOT ConveyorIO11128.xEmpty,PT:= t#3s ,Q:= m_x111271 ,ET:= m_t111271);
		IF NOT ConveyorIO11128.xEmpty AND m_x111271 THEN(*加延时刷新111261，线体第0步要延时100ms才能检测有料，*)
			ConveyorIO111271.xPutInto:=1;
		ELSIF ConveyorIO111271.xEmpty=0 THEN
			ConveyorIO111271.xPutInto:=0;
		END_IF;	

		ConveyorIO11128.xUnload:=ConveyorIO11127.xEmpty AND UConveyorio11312.iTask=2 ;
		(*至此，U4的动作全部完成*)

		(*机械手完空框回流*)
		(*12203升降控制*)
		LifterIO11203.xMDIExe:= NOT ConveyorIO11116.xError AND  NOT ConveyorIO11117.xError  AND  NOT ConveyorIO11130.xError ;
		IF ConveyorIO11117.xEmpty THEN
			LifterIO11203.iDestinationPos:=2;
		ELSE
			LifterIO11203.iDestinationPos:=1;
		END_IF;		
		ConveyorIO11116.xUnload:=ConveyorIO11116.diDesConveyor=11117 AND ConveyorIO11117.xEmpty AND  LifterIO11203.iCurrentPos=2;
		ConveyorIO11117.xUnloadCCW:=1; 
		ConveyorIO11117.xLoad:=ConveyorIO11116.xNextRun AND LifterIO11203.iCurrentPos=2;
		ConveyorIO11117.xUnload:=LifterIO11203.iCurrentPos=1 	AND ConveyorIO11130.xEmpty;
		ConveyorIO11130.xLoad:=	ConveyorIO11117.xNextRun;	
		ConveyorIO11130.xUnload:=	ConveyorIO11131.xEmpty;
		ConveyorIO11131.xLoad:=	ConveyorIO11130.xNextRun;	
		ConveyorIO11131.xUnload:=	ConveyorIO11132.xEmpty;
		ConveyorIO11132.xLoad:=	ConveyorIO11131.xNextRun;	
		ConveyorIO11132.xUnload:=	ConveyorIO11133.xEmpty;
		ConveyorIO11133.xLoad:=	ConveyorIO11132.xNextRun;	
		ConveyorIO11133.xUnload:=	ConveyorIO11134.xEmpty;
		ConveyorIO11134.xLoad:=	ConveyorIO11133.xNextRun;	
		ConveyorIO11134.xUnload:=	ConveyorIO11135.xEmpty;
		ConveyorIO11135.xLoad:=	ConveyorIO11134.xNextRun;		
		ConveyorIO11135.xUnload:=ConveyorIO11136.xEmpty;
		ConveyorIO11136.xLoad:=	ConveyorIO11135.xNextRun;	
		ConveyorIO11136.xUnload:=	ConveyorIO11137.xEmpty AND m_i11315Task=1 AND NOT  conveyorIO11137.xError; (*传递到11315了，要转方向了*)
		ConveyorIO11143.xLoad:=ConveyorIO111381.xNextRun AND m_i11315Task=1;
		CylinderIO112041.xMDIExe:=1;
		IF ConveyorIO11143.xEmpty=0 AND ConveyorIO11144.xEmpty AND CylinderIO112041.iCurrentPos=2  THEN
			CylinderIO112042.iDestinationPos:=1;
		ELSE
			CylinderIO112042.iDestinationPos:=2;
		END_IF;
		CylinderIO112042.xMDIExe:=1;
		IF D401.0 AND NOT ConveyorIO11144.xEmpty  AND CylinderIO112042.iCurrentPos=2 THEN
			CylinderIO112041.iDestinationPos:=1;
		ELSE
			CylinderIO112041.iDestinationPos:=2;
		END_IF;
			ConveyorIO11143.xUnload:=ConveyorIO11144.xEmpty AND CylinderIO112042.iCurrentPos=1;
			ConveyorIO11144.xLoad:=ConveyorIO11143.xNextRun;
			ConveyorIO11144.xUnload:=D401.0 AND CylinderIO112041.iCurrentPos=1;
			D201.0:=ConveyorIO11144.xNextRun;(*到这里运到了10那边去*)